// TIA Portal project "TIA1200_Level1" (V19)

(* hardware
DEVICE "S7-1200 station_1"  S7-1200 Station
   slot 0: "Rack_0"  S7-1200 Rack  Rack  V1.0
   slot 1: "PLC_1"  CPU 1214C DC/DC/DC  6ES7 214-1AG40-0XB0  V4.6
   slot 3: "AQ 1x12BIT_1"  AQ1 signal board  6ES7 232-4HA30-0XB0  V1.0
DEVICE "HMI_1"  KTP700 Basic PN
   slot 0: "HMI_1"  KTP700 Basic PN  6AV2 123-2GB03-0AX0  17.0.0.0
   slot 1: "HMI_RT_1"  KTP700 Basic PN  6AV2 123-2GB03-0AX0  17.0.0.0
   slot 5: "HMI_1.IE_CP_1"  PROFINET Interface  17.0.0.0
      slot 1: "PROFINET Interface_1"  PROFINET Interface
         slot 1: "Port_1"  Port
*)

// ===== PLC "PLC_1"  CPU 1214C DC/DC/DC =====

VAR_GLOBAL   // PLC tag table "Default tag table"
   "System_Byte" AT %MB1 : Byte;
   "FirstScan" AT %M1.0 : Bool;
   "DiagStatusUpdate" AT %M1.1 : Bool;
   "AlwaysTRUE" AT %M1.2 : Bool;
   "AlwaysFALSE" AT %M1.3 : Bool;
   "Clock_Byte" AT %MB0 : Byte;
   "Clock_10Hz" AT %M0.0 : Bool;
   "Clock_5Hz" AT %M0.1 : Bool;
   "Clock_2.5Hz" AT %M0.2 : Bool;
   "Clock_2Hz" AT %M0.3 : Bool;
   "Clock_1.25Hz" AT %M0.4 : Bool;
   "Clock_1Hz" AT %M0.5 : Bool;
   "Clock_0.625Hz" AT %M0.6 : Bool;
   "Clock_0.5Hz" AT %M0.7 : Bool;
END_VAR

VAR_GLOBAL   // PLC tag table "Inputs-Outputs"
   "Button OFF" AT %I0.0 : Bool;
   "Button ON" AT %I0.1 : Bool;
   "E-Stop" AT %I0.2 : Bool;
   "Cylinder A retracted" AT %I0.3 : Bool;
   "Cylinder B extended" AT %I0.4 : Bool;
   "Gripper open" AT %I0.5 : Bool;
   "Cylinder A extended" AT %I0.6 : Bool;
   "Cylinder B retracted" AT %I0.7 : Bool;
   "Button0" AT %I1.0 : Bool;
   "Button1" AT %I1.1 : Bool;
   "Button2" AT %I1.2 : Bool;
   "Button3" AT %I1.3 : Bool;
   "Button4" AT %I1.4 : Bool;
   "Button5" AT %I1.5 : Bool;
   "Retract cylinder A" AT %Q0.0 : Bool;
   "Extend cylinder B" AT %Q0.1 : Bool;
   "Close the gripper" AT %Q0.2 : Bool;
   "Extend cylinder A" AT %Q0.3 : Bool;
   "Lamp" AT %Q0.4 : Bool;
   "Retract cylinder B" AT %Q0.5 : Bool;
   "0–10V display" AT %QW80 : Int;
   "Potentiometer 1 (0–10V)" AT %IW64 : Int;
END_VAR

DATA_BLOCK "DB001_Alarms_Handling"   // DB1
{ S7_Optimized_Access := 'TRUE' }
VERSION : 0.1
   VAR
      Alarm_Active : Bool;
      Alarm_Cause : Bool;
      Auxilary0 : Bool;
   END_VAR
BEGIN
END_DATA_BLOCK

DATA_BLOCK "DB002_Auto_Cycle"   // DB2
{ S7_Optimized_Access := 'TRUE' }
VERSION : 0.1
   VAR
      Auto : Bool;
      Auxilary0 : Bool;
      Auxilary1 : Bool;
      HMI_Start : Bool;
      HMI_Stop : Bool;
   END_VAR
BEGIN
END_DATA_BLOCK

DATA_BLOCK "DB003_Calculations"   // DB3
{ S7_Optimized_Access := 'TRUE' }
VERSION : 0.1
   VAR
      Stock : Int;
      Sum : Int;
      Sum1 : Int := 50;
      Sum2 : Int := 45;
      Losses : Int := 10;
      ParDod : Int := 1;
      Auxilary0 : Bool;
   END_VAR
BEGIN
END_DATA_BLOCK

DATA_BLOCK "DB004_Labeler_Control"   // DB4
{ S7_Optimized_Access := 'TRUE' }
VERSION : 0.1
   VAR
      Label_Roll_Length : Int := 5000;
      Current_Label_Roll_Length : Int;
      Label_Length : Int := 250;
      Labels_Counter : Int;
      Label_Rolls_Counter : Int;
      Number_of_Labels_Remaining : Int;
      Unwind_Permission : Bool;
      Auxilary0 : Bool;
      Auxilary1 : Bool;
   END_VAR
BEGIN
END_DATA_BLOCK

DATA_BLOCK "DB007_Pulse_Generator"   // DB7
{ S7_Optimized_Access := 'TRUE' }
VERSION : 0.1
   VAR
      Generator_Status : Bool;
      Time_ON : Time := T#2s;
      Time_OFF : Time := T#2s;
   END_VAR
BEGIN
END_DATA_BLOCK

DATA_BLOCK "DB011_Motor_With_Cooling"   // DB11
{ S7_Optimized_Access := 'TRUE' }
VERSION : 0.1
   VAR
      "E-Stop Alarm" : Bool;
      Auxilary0 : Bool;
   END_VAR
BEGIN
END_DATA_BLOCK

DATA_BLOCK "DB012_Cylinder_Timout"   // DB13
{ S7_Optimized_Access := 'TRUE' }
VERSION : 0.1
   VAR
      "Timout Alarm" : Bool;
      Auxilary0 : Bool;
   END_VAR
BEGIN
END_DATA_BLOCK

DATA_BLOCK "DB015_Three_Production_Lines"   // DB16
{ S7_Optimized_Access := 'TRUE' }
VERSION : 0.1
   VAR
      "Line#1 Qty" : UDInt;
      "Line#2 Qty" : UDInt;
      "Line#3 Qty" : UDInt;
      "Line#1 UnitPrice" : Int := 4;
      "Line#2 UnitPrice" : Int := 3;
      "Line#3 UnitPrice" : Int := 39;
      "Total Profit" : UDInt;
      Auxilary0 : Bool;
      Auxilary1 : Bool;
      Auxilary2 : Bool;
   END_VAR
BEGIN
END_DATA_BLOCK

DATA_BLOCK "DB017_Packaging_Control"   // DB18
{ S7_Optimized_Access := 'TRUE' }
VERSION : 0.1
   VAR
      "Next Row" : Bool;
      "Next Box" : Bool;
      "Boxes Total Qty" : UDInt;
      "Box Fill Count" : Int;
   END_VAR
BEGIN
END_DATA_BLOCK

// folder: System blocks/Program resources

DATA_BLOCK "DB005_Buffer_Filling"   // DB5
{ S7_Optimized_Access := 'TRUE' }
AUTHOR : Simatic
FAMILY : IEC
NAME : CNTR
VERSION : 1.0
// stored: InstanceOfName IEC_COUNTER
"IEC_COUNTER"
BEGIN
END_DATA_BLOCK

DATA_BLOCK "DB006_Lift_Sequence"   // DB6
{ S7_Optimized_Access := 'TRUE' }
AUTHOR : Simatic
FAMILY : IEC
NAME : CNTR
VERSION : 1.0
// stored: InstanceOfName IEC_COUNTER
"IEC_COUNTER"
BEGIN
END_DATA_BLOCK

DATA_BLOCK "DB008_PulseGenerator_TimerOFF"   // DB8
{ S7_Optimized_Access := 'TRUE' }
AUTHOR : Simatic
FAMILY : IEC
NAME : IEC_TMR
VERSION : 1.0
// stored: InstanceOfName IEC_TIMER
"IEC_TIMER"
BEGIN
END_DATA_BLOCK

DATA_BLOCK "DB008_PulseGenerator_TimerON"   // DB9
{ S7_Optimized_Access := 'TRUE' }
AUTHOR : Simatic
FAMILY : IEC
NAME : IEC_TMR
VERSION : 1.0
// stored: InstanceOfName IEC_TIMER
"IEC_TIMER"
BEGIN
END_DATA_BLOCK

DATA_BLOCK "DB009_MotorWithCooling_TON"   // DB10
{ S7_Optimized_Access := 'TRUE' }
AUTHOR : Simatic
FAMILY : IEC
NAME : IEC_TMR
VERSION : 1.0
// stored: InstanceOfName IEC_TIMER
"IEC_TIMER"
BEGIN
END_DATA_BLOCK

DATA_BLOCK "DB010_MotorWithCooling_TOF"   // DB12
{ S7_Optimized_Access := 'TRUE' }
AUTHOR : Simatic
FAMILY : IEC
NAME : IEC_TMR
VERSION : 1.0
// stored: InstanceOfName IEC_TIMER
"IEC_TIMER"
BEGIN
END_DATA_BLOCK

DATA_BLOCK "DB013_CylinderTimeout_Extend_TON"   // DB14
{ S7_Optimized_Access := 'TRUE' }
AUTHOR : Simatic
FAMILY : IEC
NAME : IEC_TMR
VERSION : 1.0
// stored: InstanceOfName IEC_TIMER
"IEC_TIMER"
BEGIN
END_DATA_BLOCK

DATA_BLOCK "DB014_CylinderTimeout_Retract_TON"   // DB15
{ S7_Optimized_Access := 'TRUE' }
AUTHOR : Simatic
FAMILY : IEC
NAME : IEC_TMR
VERSION : 1.0
// stored: InstanceOfName IEC_TIMER
"IEC_TIMER"
BEGIN
END_DATA_BLOCK

DATA_BLOCK "DB016_PackagingControl_Units"   // DB17
{ S7_Optimized_Access := 'TRUE' }
AUTHOR : Simatic
FAMILY : IEC
NAME : CNTR
VERSION : 1.0
// stored: InstanceOfName IEC_COUNTER
"IEC_COUNTER"
BEGIN
END_DATA_BLOCK

DATA_BLOCK "DB018_PackagingControl_Row"   // DB19
{ S7_Optimized_Access := 'TRUE' }
AUTHOR : Simatic
FAMILY : IEC
NAME : CNTR
VERSION : 1.0
// stored: InstanceOfName IEC_COUNTER
"IEC_COUNTER"
BEGIN
END_DATA_BLOCK

DATA_BLOCK "DB019_PacakagingControl_BoxFillCnt"   // DB20
{ S7_Optimized_Access := 'TRUE' }
AUTHOR : Simatic
FAMILY : IEC
NAME : CNTR
VERSION : 1.0
// stored: InstanceOfName IEC_COUNTER
"IEC_COUNTER"
BEGIN
END_DATA_BLOCK

// folder: (top level)

FUNCTION "FC001_Close_Gripper" : Void   // FC1, LAD
{ S7_Optimized_Access := 'TRUE' }
VERSION : 0.1
BEGIN

REGION Network 1: Close Gripper Logic
   // Pressing the green button I0.1 causes the gripper to close on output Q0.2
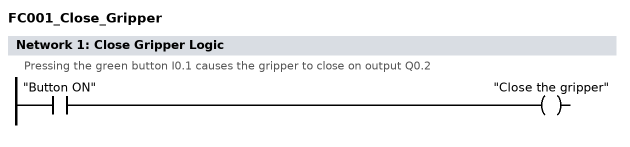
   RUNG wire#powerrail
      Contact( "Button ON" )
      Coil( "Close the gripper" )
   END_RUNG
   // the same network as SCL:
   "Close the gripper" := "Button ON";
END_REGION
END_FUNCTION

FUNCTION "FC002_PusherA_Operation" : Void   // FC2, LAD
{ S7_Optimized_Access := 'TRUE' }
VERSION : 0.1
BEGIN

REGION Network 1: Cylinder A Control Logic
   // Pressing button I0.1 extends cylinder A (Q0.3). Releasing the button and activating I0.0 retracts cylinder A (Q0.0)
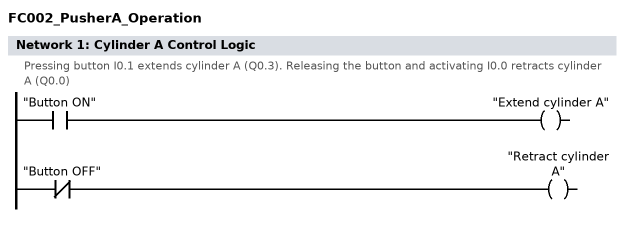
   RUNG wire#powerrail
      Contact( "Button ON" )
      Coil( "Extend cylinder A" )
   END_RUNG
   RUNG wire#powerrail
      I_Contact( "Button OFF" )
      Coil( "Retract cylinder A" )
   END_RUNG
   // the same network as SCL:
   "Extend cylinder A" := "Button ON";
   "Retract cylinder A" := NOT "Button OFF";
END_REGION
END_FUNCTION

FUNCTION "FC003_PusherB_Operation" : Void   // FC3, LAD
{ S7_Optimized_Access := 'TRUE' }
VERSION : 0.1
BEGIN

REGION Network 1: Cylinder B Control Logic
   // Pressing the silver switch I1.3 extends cylinder B on Q0.1. Pressing the silver switch I1.4 retracts cylinder B on Q0.5
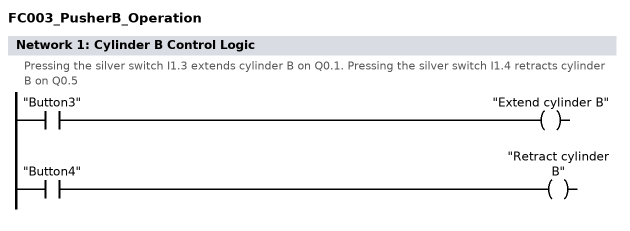
   RUNG wire#powerrail
      Contact( "Button3" )
      Coil( "Extend cylinder B" )
   END_RUNG
   RUNG wire#powerrail
      Contact( "Button4" )
      Coil( "Retract cylinder B" )
   END_RUNG
   // the same network as SCL:
   "Extend cylinder B" := "Button3";
   "Retract cylinder B" := "Button4";
END_REGION
END_FUNCTION

FUNCTION "FC001_Close_Gripper#2" : Void   // FC4, LAD
{ S7_Optimized_Access := 'TRUE' }
VERSION : 0.1
BEGIN

REGION Network 1: Close Gripper Logic
   // The gripper closes when the green button is pressed and both cylinder A and cylinder B are in the extended position
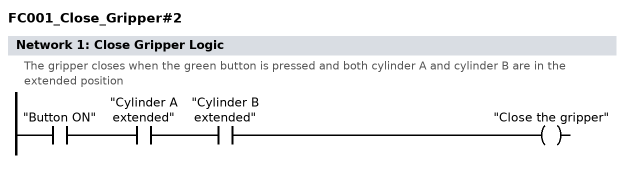
   RUNG wire#powerrail
      Contact( "Button ON" )
      Contact( "Cylinder A extended" )
      Contact( "Cylinder B extended" )
      Coil( "Close the gripper" )
   END_RUNG
   // the same network as SCL:
   "Close the gripper" := "Button ON" AND "Cylinder A extended" AND "Cylinder B extended";
END_REGION
END_FUNCTION

FUNCTION "FC002_PusherA_Operation_Safty" : Void   // FC5, LAD
{ S7_Optimized_Access := 'TRUE' }
VERSION : 0.1
BEGIN

REGION Network 1: Cylinder A Control Logic + Safty
   // Pressing button I0.1 extends cylinder A (Q0.3), but the output is disabled when the upper position sensor I0.6 is activated. 
   // Pressing button I0.0 retracts cylinder A (Q0.0), but the output is disabled when the lower position sensor I0.3 is activated. 
   // Additionally, pressing the emergency stop button I0.2 disables all motion and prevents the pusher from operating.
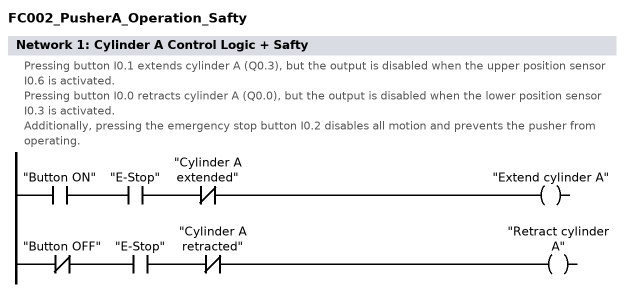
   RUNG wire#powerrail
      Contact( "Button ON" )
      Contact( "E-Stop" )
      I_Contact( "Cylinder A extended" )
      Coil( "Extend cylinder A" )
   END_RUNG
   RUNG wire#powerrail
      I_Contact( "Button OFF" )
      Contact( "E-Stop" )
      I_Contact( "Cylinder A retracted" )
      Coil( "Retract cylinder A" )
   END_RUNG
   // the same network as SCL:
   "Extend cylinder A" := "Button ON" AND "E-Stop" AND NOT "Cylinder A extended";
   "Retract cylinder A" := NOT "Button OFF" AND "E-Stop" AND NOT "Cylinder A retracted";
END_REGION
END_FUNCTION

FUNCTION "FC002_PusherA_Operation_Signalling" : Void   // FC6, LAD
{ S7_Optimized_Access := 'TRUE' }
VERSION : 0.1
BEGIN

REGION Network 1: Cylinder A Control Logic + Safty
   // Pressing button I0.1 extends cylinder A (Q0.3), but the output is disabled when the upper position sensor I0.6 is activated. 
   // Pressing button I0.0 retracts cylinder A (Q0.0), but the output is disabled when the lower position sensor I0.3 is activated. 
   // Additionally, pressing the emergency stop button I0.2 disables all motion and prevents the pusher from operating.
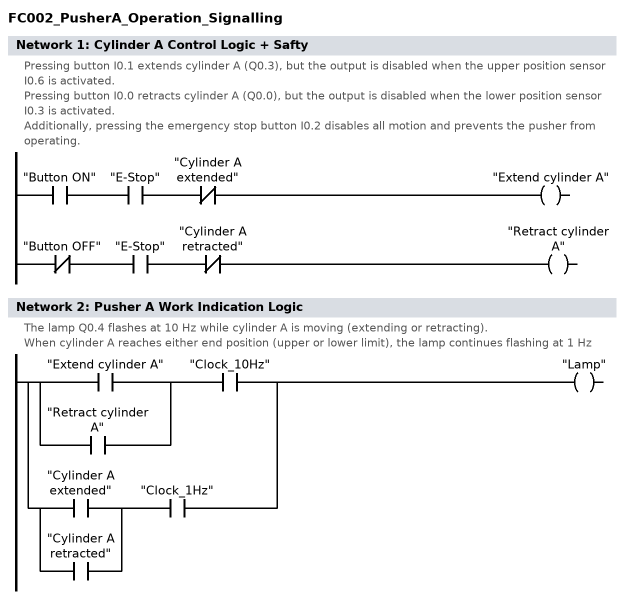
   RUNG wire#powerrail
      Contact( "Button ON" )
      Contact( "E-Stop" )
      I_Contact( "Cylinder A extended" )
      Coil( "Extend cylinder A" )
   END_RUNG
   RUNG wire#powerrail
      I_Contact( "Button OFF" )
      Contact( "E-Stop" )
      I_Contact( "Cylinder A retracted" )
      Coil( "Retract cylinder A" )
   END_RUNG
   // the same network as SCL:
   "Extend cylinder A" := "Button ON" AND "E-Stop" AND NOT "Cylinder A extended";
   "Retract cylinder A" := NOT "Button OFF" AND "E-Stop" AND NOT "Cylinder A retracted";
END_REGION

REGION Network 2: Pusher A Work Indication Logic
   // The lamp Q0.4 flashes at 10 Hz while cylinder A is moving (extending or retracting). 
   // When cylinder A reaches either end position (upper or lower limit), the lamp continues flashing at 1 Hz
   RUNG wire#powerrail
      Contact( "Extend cylinder A" )
      wire#w1
      Contact( "Clock_10Hz" )
      wire#w2
      Coil( "Lamp" )
   END_RUNG
   RUNG wire#powerrail
      Contact( "Retract cylinder A" )
   END_RUNG wire#w1
   RUNG wire#powerrail
      Contact( "Cylinder A extended" )
      wire#w3
      Contact( "Clock_1Hz" )
   END_RUNG wire#w2
   RUNG wire#powerrail
      Contact( "Cylinder A retracted" )
   END_RUNG wire#w3
   // the same network as SCL:
   "Lamp" := (("Extend cylinder A" OR "Retract cylinder A") AND "Clock_10Hz") OR (("Cylinder A extended" OR "Cylinder A retracted") AND "Clock_1Hz");
END_REGION
END_FUNCTION

FUNCTION "FC004_EndPosition" : Void   // FC7, LAD
{ S7_Optimized_Access := 'TRUE' }
VERSION : 0.1
BEGIN

REGION Network 1: Extend Cylinder A Logic
   // Button ON extends cylinder A until the upper limit I0.6 is reached
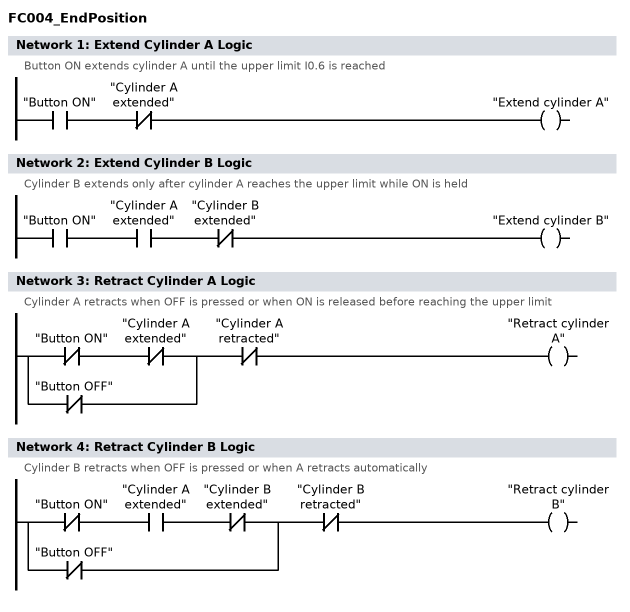
   RUNG wire#powerrail
      Contact( "Button ON" )
      I_Contact( "Cylinder A extended" )
      Coil( "Extend cylinder A" )
   END_RUNG
   // the same network as SCL:
   "Extend cylinder A" := "Button ON" AND NOT "Cylinder A extended";
END_REGION

REGION Network 2: Extend Cylinder B Logic
   // Cylinder B extends only after cylinder A reaches the upper limit while ON is held
   RUNG wire#powerrail
      Contact( "Button ON" )
      Contact( "Cylinder A extended" )
      I_Contact( "Cylinder B extended" )
      Coil( "Extend cylinder B" )
   END_RUNG
   // the same network as SCL:
   "Extend cylinder B" := "Button ON" AND "Cylinder A extended" AND NOT "Cylinder B extended";
END_REGION

REGION Network 3: Retract Cylinder A Logic
   // Cylinder A retracts when OFF is pressed or when ON is released before reaching the upper limit
   RUNG wire#powerrail
      I_Contact( "Button ON" )
      I_Contact( "Cylinder A extended" )
      wire#w1
      I_Contact( "Cylinder A retracted" )
      Coil( "Retract cylinder A" )
   END_RUNG
   RUNG wire#powerrail
      I_Contact( "Button OFF" )
   END_RUNG wire#w1
   // the same network as SCL:
   "Retract cylinder A" := ((NOT "Button ON" AND NOT "Cylinder A extended") OR NOT "Button OFF") AND NOT "Cylinder A retracted";
END_REGION

REGION Network 4: Retract Cylinder B Logic
   // Cylinder B retracts when OFF is pressed or when A retracts automatically
   RUNG wire#powerrail
      I_Contact( "Button ON" )
      Contact( "Cylinder A extended" )
      I_Contact( "Cylinder B extended" )
      wire#w1
      I_Contact( "Cylinder B retracted" )
      Coil( "Retract cylinder B" )
   END_RUNG
   RUNG wire#powerrail
      I_Contact( "Button OFF" )
   END_RUNG wire#w1
   // the same network as SCL:
   "Retract cylinder B" := ((NOT "Button ON" AND "Cylinder A extended" AND NOT "Cylinder B extended") OR NOT "Button OFF") AND NOT "Cylinder B retracted";
END_REGION
END_FUNCTION

FUNCTION "FC005_Element_Position_Control" : Void   // FC8, LAD
{ S7_Optimized_Access := 'TRUE' }
VERSION : 0.1
BEGIN

REGION Network 1: Element Position Control Logic
   // Lamp Q0.4 is ON when all sensors are active, flashes at 2 Hz when only one sensor is missing, and remains OFF when at most one sensor is active
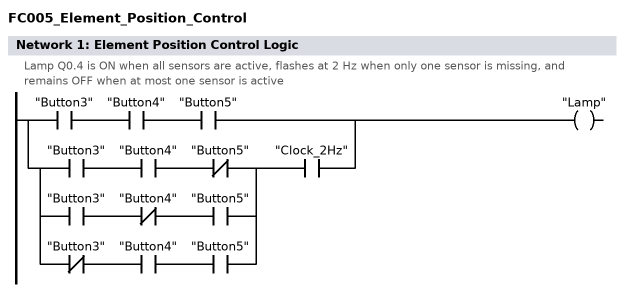
   RUNG wire#powerrail
      Contact( "Button3" )
      Contact( "Button4" )
      Contact( "Button5" )
      wire#w1
      Coil( "Lamp" )
   END_RUNG
   RUNG wire#powerrail
      Contact( "Button3" )
      Contact( "Button4" )
      I_Contact( "Button5" )
      wire#w2
      Contact( "Clock_2Hz" )
   END_RUNG wire#w1
   RUNG wire#powerrail
      Contact( "Button3" )
      I_Contact( "Button4" )
      Contact( "Button5" )
   END_RUNG wire#w2
   RUNG wire#powerrail
      I_Contact( "Button3" )
      Contact( "Button4" )
      Contact( "Button5" )
   END_RUNG wire#w2
   // the same network as SCL:
   "Lamp" := ("Button3" AND "Button4" AND "Button5") OR ((("Button3" AND "Button4" AND NOT "Button5") OR ("Button3" AND NOT "Button4" AND "Button5") OR (NOT "Button3" AND "Button4" AND "Button5")) AND "Clock_2Hz");
END_REGION
END_FUNCTION

FUNCTION "FC006_Robot_Gripper_Control" : Void   // FC9, LAD
{ S7_Optimized_Access := 'TRUE' }
VERSION : 0.1
BEGIN

REGION Network 1: Gripper Open / Close Logic
   // Pressing ON closes the gripper. Pressing OFF (NC) closes the gripper
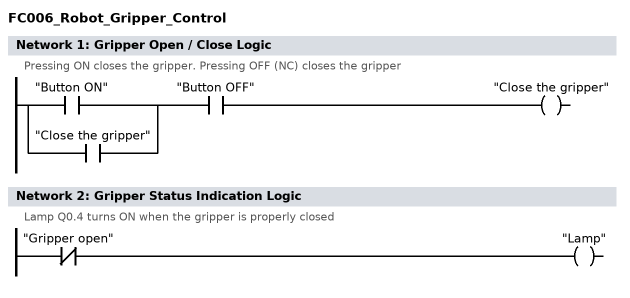
   RUNG wire#powerrail
      Contact( "Button ON" )
      wire#w1
      Contact( "Button OFF" )
      Coil( "Close the gripper" )
   END_RUNG
   RUNG wire#powerrail
      Contact( "Close the gripper" )
   END_RUNG wire#w1
   // the same network as SCL:
   "Close the gripper" := ("Button ON" OR "Close the gripper") AND "Button OFF";
END_REGION

REGION Network 2: Gripper Status Indication Logic
   // Lamp Q0.4 turns ON when the gripper is properly closed
   RUNG wire#powerrail
      I_Contact( "Gripper open" )
      Coil( "Lamp" )
   END_RUNG
   // the same network as SCL:
   "Lamp" := NOT "Gripper open";
END_REGION
END_FUNCTION

FUNCTION "FC006_Robot_Gripper_Control#2" : Void   // FC10, LAD
{ S7_Optimized_Access := 'TRUE' }
VERSION : 0.1
BEGIN

REGION Network 1: Gripper Open / Close Logic
   // Pressing ON closes the gripper. Pressing OFF (NC) closes the gripper with Set/Reset block
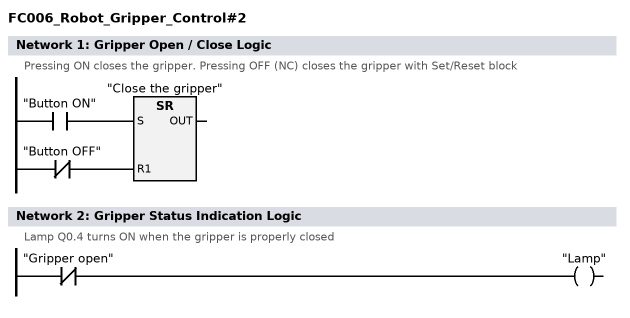
   RUNG wire#powerrail
      Contact( "Button ON" )
      S_SR(operand := "Close the gripper", r1 := wire#w1)
   END_RUNG
   RUNG wire#powerrail
      I_Contact( "Button OFF" )
   END_RUNG wire#w1
   // the same network as SCL:
   IF "Button ON" THEN
       "Close the gripper" := TRUE;   // SR flip-flop
   END_IF;
   IF NOT "Button OFF" THEN "Close the gripper" := FALSE; END_IF;
END_REGION

REGION Network 2: Gripper Status Indication Logic
   // Lamp Q0.4 turns ON when the gripper is properly closed
   RUNG wire#powerrail
      I_Contact( "Gripper open" )
      Coil( "Lamp" )
   END_RUNG
   // the same network as SCL:
   "Lamp" := NOT "Gripper open";
END_REGION
END_FUNCTION

FUNCTION "FC007_Pneumatic_Lift" : Void   // FC11, LAD
{ S7_Optimized_Access := 'TRUE' }
VERSION : 0.1
BEGIN

REGION Network 1: Lift Extend Logic
   // Switch I1.3 extends cylinder A on Q0.3; the output is cut off at the upper limit I0.6
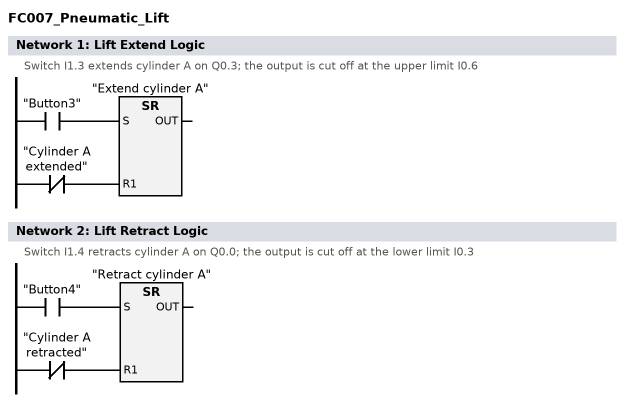
   RUNG wire#powerrail
      Contact( "Button3" )
      S_SR(operand := "Extend cylinder A", r1 := wire#w1)
   END_RUNG
   RUNG wire#powerrail
      I_Contact( "Cylinder A extended" )
   END_RUNG wire#w1
   // the same network as SCL:
   IF "Button3" THEN
       "Extend cylinder A" := TRUE;   // SR flip-flop
   END_IF;
   IF NOT "Cylinder A extended" THEN "Extend cylinder A" := FALSE; END_IF;
END_REGION

REGION Network 2: Lift Retract Logic
   // Switch I1.4 retracts cylinder A on Q0.0; the output is cut off at the lower limit I0.3
   RUNG wire#powerrail
      Contact( "Button4" )
      S_SR(operand := "Retract cylinder A", r1 := wire#w1)
   END_RUNG
   RUNG wire#powerrail
      I_Contact( "Cylinder A retracted" )
   END_RUNG wire#w1
   // the same network as SCL:
   IF "Button4" THEN
       "Retract cylinder A" := TRUE;   // SR flip-flop
   END_IF;
   IF NOT "Cylinder A retracted" THEN "Retract cylinder A" := FALSE; END_IF;
END_REGION
END_FUNCTION

FUNCTION "FC008_Alarms_Handling" : Void   // FC12, LAD
{ S7_Optimized_Access := 'TRUE' }
VERSION : 0.1
   VAR_TEMP   // added for the SCL form of the ladder/FBD networks
      _w1 : Bool;
   END_VAR
BEGIN

REGION Network 1: Alarm Cause Evaluation
   // Evaluate alarm cause. Normal operating state:
   // 
   // I1.0=1 (Fuse), I1.1=1 (Motor temperature), I1.2=0 (Pusher interlock), I1.3=0 (Pressure OK).
   // Set Alarm_Cause when any input deviates from its normal state
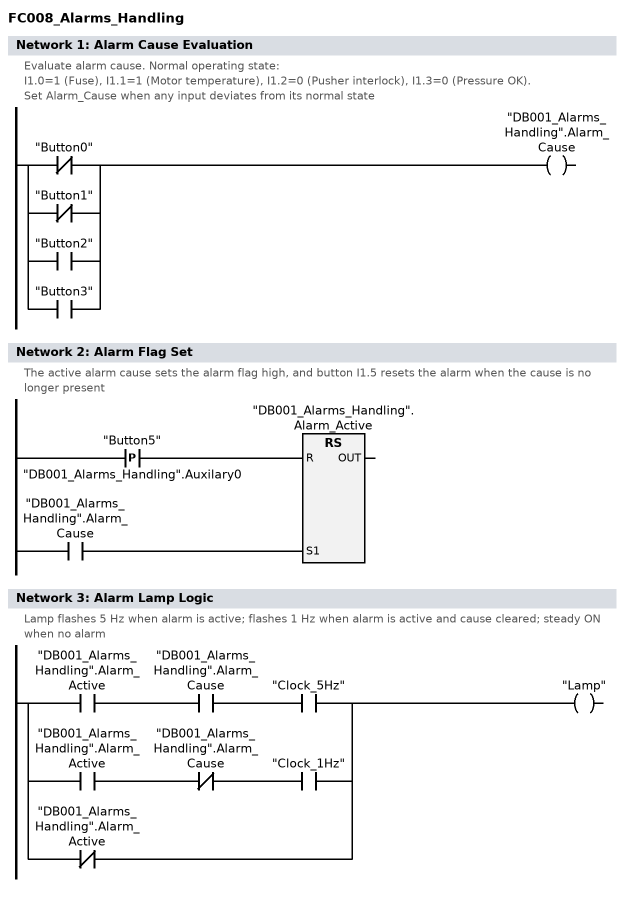
   RUNG wire#powerrail
      I_Contact( "Button0" )
      wire#w1
      Coil( "DB001_Alarms_Handling".Alarm_Cause )
   END_RUNG
   RUNG wire#powerrail
      I_Contact( "Button1" )
   END_RUNG wire#w1
   RUNG wire#powerrail
      Contact( "Button2" )
   END_RUNG wire#w1
   RUNG wire#powerrail
      Contact( "Button3" )
   END_RUNG wire#w1
   // the same network as SCL:
   "DB001_Alarms_Handling".Alarm_Cause := NOT "Button0" OR NOT "Button1" OR "Button2" OR "Button3";
END_REGION

REGION Network 2: Alarm Flag Set
   // The active alarm cause sets the alarm flag high, and button I1.5 resets the alarm when the cause is no longer present
   RUNG wire#powerrail
      P_Contact(operand := "Button5", bit := "DB001_Alarms_Handling".Auxilary0)
      S_RS(operand := "DB001_Alarms_Handling".Alarm_Active, s1 := wire#w1)
   END_RUNG
   RUNG wire#powerrail
      Contact( "DB001_Alarms_Handling".Alarm_Cause )
   END_RUNG wire#w1
   // the same network as SCL:
   #_w1 := "Button5" AND NOT "DB001_Alarms_Handling".Auxilary0;   // rising edge of "Button5"
   "DB001_Alarms_Handling".Auxilary0 := "Button5";
   IF #_w1 THEN
       "DB001_Alarms_Handling".Alarm_Active := FALSE;   // RS flip-flop
   END_IF;
   IF "DB001_Alarms_Handling".Alarm_Cause THEN "DB001_Alarms_Handling".Alarm_Active := TRUE; END_IF;
END_REGION

REGION Network 3: Alarm Lamp Logic
   // Lamp flashes 5 Hz when alarm is active; flashes 1 Hz when alarm is active and cause cleared; steady ON when no alarm
   RUNG wire#powerrail
      Contact( "DB001_Alarms_Handling".Alarm_Active )
      Contact( "DB001_Alarms_Handling".Alarm_Cause )
      Contact( "Clock_5Hz" )
      wire#w1
      Coil( "Lamp" )
   END_RUNG
   RUNG wire#powerrail
      Contact( "DB001_Alarms_Handling".Alarm_Active )
      I_Contact( "DB001_Alarms_Handling".Alarm_Cause )
      Contact( "Clock_1Hz" )
   END_RUNG wire#w1
   RUNG wire#powerrail
      I_Contact( "DB001_Alarms_Handling".Alarm_Active )
   END_RUNG wire#w1
   // the same network as SCL:
   "Lamp" := ("DB001_Alarms_Handling".Alarm_Active AND "DB001_Alarms_Handling".Alarm_Cause AND "Clock_5Hz") OR ("DB001_Alarms_Handling".Alarm_Active AND NOT "DB001_Alarms_Handling".Alarm_Cause AND "Clock_1Hz") OR NOT "DB001_Alarms_Handling".Alarm_Active;
END_REGION
END_FUNCTION

FUNCTION "FC009_Auto_Cycle" : Void   // FC13, LAD
{ S7_Optimized_Access := 'TRUE' }
VERSION : 0.1
   VAR_TEMP   // added for the SCL form of the ladder/FBD networks
      _w1 : Bool;
   END_VAR
BEGIN

REGION Network 1: Automatic Cycle Start Logic
   // Start auto cycle with button ON or START CYCLE on HMI; stop cycle after button OFF or HMI STOP CYCLE
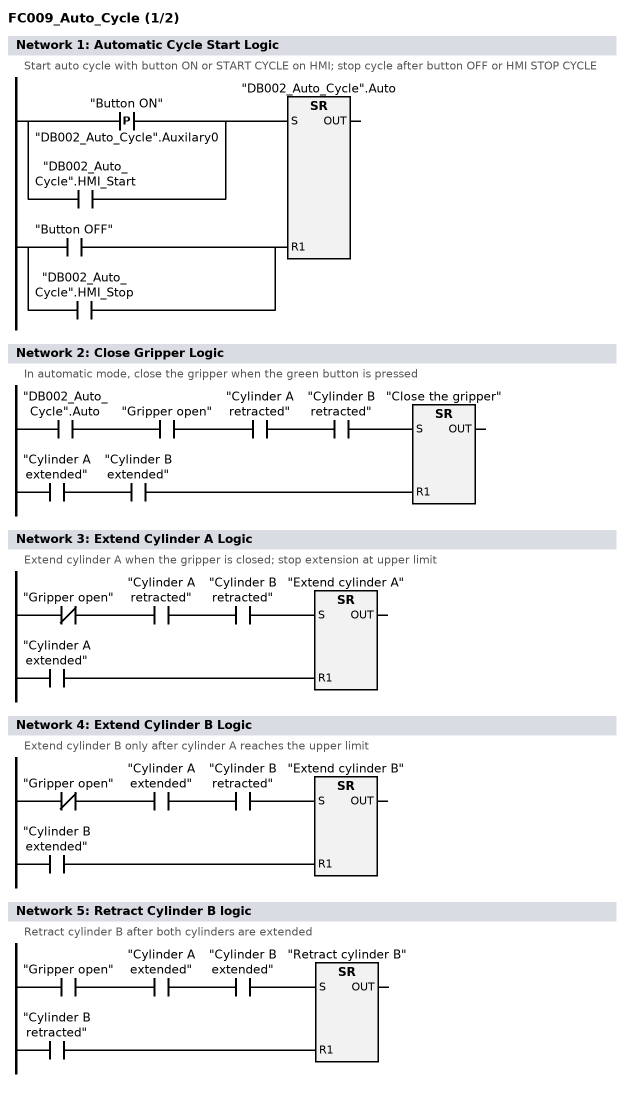
   RUNG wire#powerrail
      P_Contact(operand := "Button ON", bit := "DB002_Auto_Cycle".Auxilary0)
      wire#w1
      S_SR(operand := "DB002_Auto_Cycle".Auto, r1 := wire#w2)
   END_RUNG
   RUNG wire#powerrail
      Contact( "DB002_Auto_Cycle".HMI_Start )
   END_RUNG wire#w1
   RUNG wire#powerrail
      Contact( "Button OFF" )
   END_RUNG wire#w2
   RUNG wire#powerrail
      Contact( "DB002_Auto_Cycle".HMI_Stop )
   END_RUNG wire#w2
   // the same network as SCL:
   #_w1 := "Button ON" AND NOT "DB002_Auto_Cycle".Auxilary0;   // rising edge of "Button ON"
   "DB002_Auto_Cycle".Auxilary0 := "Button ON";
   IF #_w1 OR "DB002_Auto_Cycle".HMI_Start THEN
       "DB002_Auto_Cycle".Auto := TRUE;   // SR flip-flop
   END_IF;
   IF "Button OFF" OR "DB002_Auto_Cycle".HMI_Stop THEN "DB002_Auto_Cycle".Auto := FALSE; END_IF;
END_REGION

REGION Network 2: Close Gripper Logic
   // In automatic mode, close the gripper when the green button is pressed
   RUNG wire#powerrail
      Contact( "DB002_Auto_Cycle".Auto )
      Contact( "Gripper open" )
      Contact( "Cylinder A retracted" )
      Contact( "Cylinder B retracted" )
      S_SR(operand := "Close the gripper", r1 := wire#w1)
   END_RUNG
   RUNG wire#powerrail
      Contact( "Cylinder A extended" )
      Contact( "Cylinder B extended" )
   END_RUNG wire#w1
   // the same network as SCL:
   IF "DB002_Auto_Cycle".Auto AND "Gripper open" AND "Cylinder A retracted" AND "Cylinder B retracted" THEN
       "Close the gripper" := TRUE;   // SR flip-flop
   END_IF;
   IF "Cylinder A extended" AND "Cylinder B extended" THEN "Close the gripper" := FALSE; END_IF;
END_REGION

REGION Network 3: Extend Cylinder A Logic
   // Extend cylinder A when the gripper is closed; stop extension at upper limit
   RUNG wire#powerrail
      I_Contact( "Gripper open" )
      Contact( "Cylinder A retracted" )
      Contact( "Cylinder B retracted" )
      S_SR(operand := "Extend cylinder A", r1 := wire#w1)
   END_RUNG
   RUNG wire#powerrail
      Contact( "Cylinder A extended" )
   END_RUNG wire#w1
   // the same network as SCL:
   IF NOT "Gripper open" AND "Cylinder A retracted" AND "Cylinder B retracted" THEN
       "Extend cylinder A" := TRUE;   // SR flip-flop
   END_IF;
   IF "Cylinder A extended" THEN "Extend cylinder A" := FALSE; END_IF;
END_REGION

REGION Network 4: Extend Cylinder B Logic
   // Extend cylinder B only after cylinder A reaches the upper limit
   RUNG wire#powerrail
      I_Contact( "Gripper open" )
      Contact( "Cylinder A extended" )
      Contact( "Cylinder B retracted" )
      S_SR(operand := "Extend cylinder B", r1 := wire#w1)
   END_RUNG
   RUNG wire#powerrail
      Contact( "Cylinder B extended" )
   END_RUNG wire#w1
   // the same network as SCL:
   IF NOT "Gripper open" AND "Cylinder A extended" AND "Cylinder B retracted" THEN
       "Extend cylinder B" := TRUE;   // SR flip-flop
   END_IF;
   IF "Cylinder B extended" THEN "Extend cylinder B" := FALSE; END_IF;
END_REGION
